// TIA Portal project "Lagerregal_4" (V20) (continued)
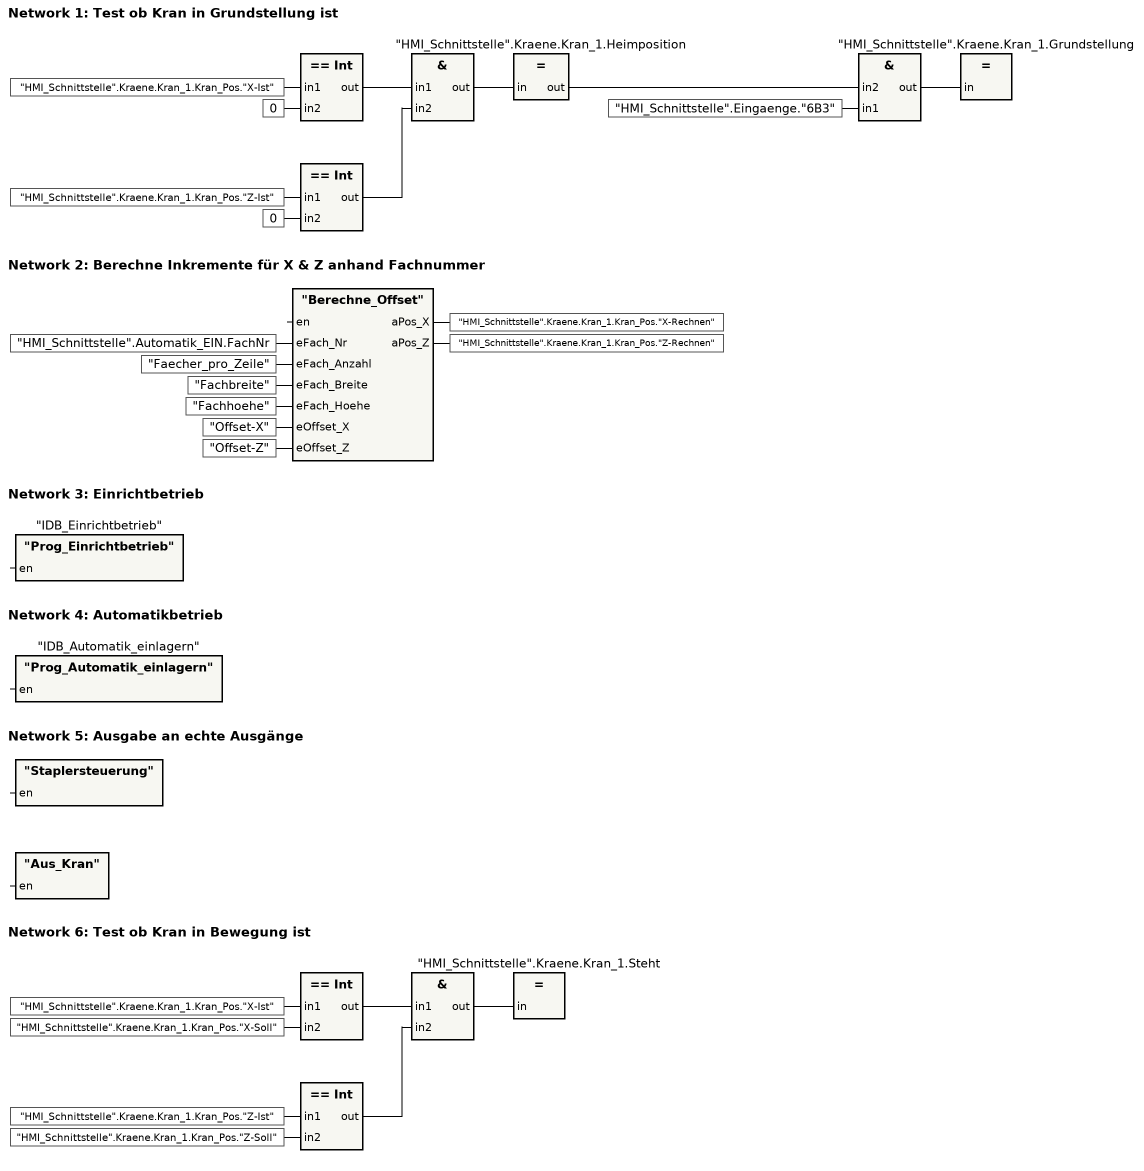
   "HMI_Schnittstelle".Kraene.Kran_1.Heimposition := ("HMI_Schnittstelle".Kraene.Kran_1.Kran_Pos."X-Ist" = 0) AND ("HMI_Schnittstelle".Kraene.Kran_1.Kran_Pos."Z-Ist" = 0);
   "HMI_Schnittstelle".Kraene.Kran_1.Grundstellung := "HMI_Schnittstelle".Kraene.Kran_1.Heimposition AND "HMI_Schnittstelle".Eingaenge."6B3";
END_REGION

REGION Network 2: Berechne Inkremente für X & Z anhand Fachnummer
   "Berechne_Offset"(eFach_Nr := "HMI_Schnittstelle".Automatik_EIN.FachNr,
                     eFach_Anzahl := "Faecher_pro_Zeile",
                     eFach_Breite := "Fachbreite",
                     eFach_Hoehe := "Fachhoehe",
                     eOffset_X := "Offset-X",
                     eOffset_Z := "Offset-Z",
                     aPos_X => "HMI_Schnittstelle".Kraene.Kran_1.Kran_Pos."X-Rechnen",
                     aPos_Z => "HMI_Schnittstelle".Kraene.Kran_1.Kran_Pos."Z-Rechnen");
END_REGION

REGION Network 3: Einrichtbetrieb
   "IDB_Einrichtbetrieb"();   // "Prog_Einrichtbetrieb"
END_REGION

REGION Network 4: Automatikbetrieb
   "IDB_Automatik_einlagern"();   // "Prog_Automatik_einlagern"
END_REGION

REGION Network 5: Ausgabe an echte Ausgänge
   "Staplersteuerung"();
   "Aus_Kran"();
END_REGION

REGION Network 6: Test ob Kran in Bewegung ist
   "HMI_Schnittstelle".Kraene.Kran_1.Steht := ("HMI_Schnittstelle".Kraene.Kran_1.Kran_Pos."X-Ist" = "HMI_Schnittstelle".Kraene.Kran_1.Kran_Pos."X-Soll") AND ("HMI_Schnittstelle".Kraene.Kran_1.Kran_Pos."Z-Ist" = "HMI_Schnittstelle".Kraene.Kran_1.Kran_Pos."Z-Soll");
END_REGION
END_ORGANIZATION_BLOCK

// folder: Bandsteuerung

FUNCTION_BLOCK "Ein_Baender"   // FB20, FBD
{ S7_Optimized_Access := 'TRUE' }
VERSION : 0.1
BEGIN

REGION Network 1 (SCL): Sensoren Einlass
   "HMI_Schnittstelle".Eingaenge."1B1" := NOT "1B1";
   "HMI_Schnittstelle".Eingaenge."1B2" := NOT "1B2";
   "HMI_Schnittstelle".Eingaenge."2B1" := NOT "2B1";
   "HMI_Schnittstelle".Eingaenge."2B2" := NOT "2B2";
   "HMI_Schnittstelle".Eingaenge."3B1" := NOT "3B1";
END_REGION

REGION Network 2 (SCL): Sensoren Auslass
   "HMI_Schnittstelle".Eingaenge."4B1" := NOT "4B1";
   "HMI_Schnittstelle".Eingaenge."5B1" := NOT "5B1";
END_REGION
END_FUNCTION_BLOCK

FUNCTION_BLOCK "Bandsteuerung"   // FB21, FBD
{ S7_Optimized_Access := 'TRUE' }
VERSION : 0.1
   VAR
      RTRIG_Palette_geladen : R_TRIG;
      FTRIG_MDB_1B2 : F_TRIG;
      FTRIG_MDB_2B1 : F_TRIG;
      FTRIG_MDB_2B2 : F_TRIG;
      FTRIG_MDB_5B1 : F_TRIG;
      Band_belegt : Bool;
   END_VAR
BEGIN

REGION Network 1 (SCL): Flankenabfragen
   #RTRIG_Palette_geladen(CLK:="HMI_Schnittstelle".Automatik_EIN.Schrittnummer = 5);
   #FTRIG_MDB_1B2(CLK:="HMI_Schnittstelle".Eingaenge."1B2");
   #FTRIG_MDB_2B1(CLK := "HMI_Schnittstelle".Eingaenge."2B1");
   #FTRIG_MDB_2B2(CLK := "HMI_Schnittstelle".Eingaenge."2B2");
   #FTRIG_MDB_5B1(CLK := "HMI_Schnittstelle".Eingaenge."5B1");
END_REGION

REGION Network 2: Einlasssteuerung
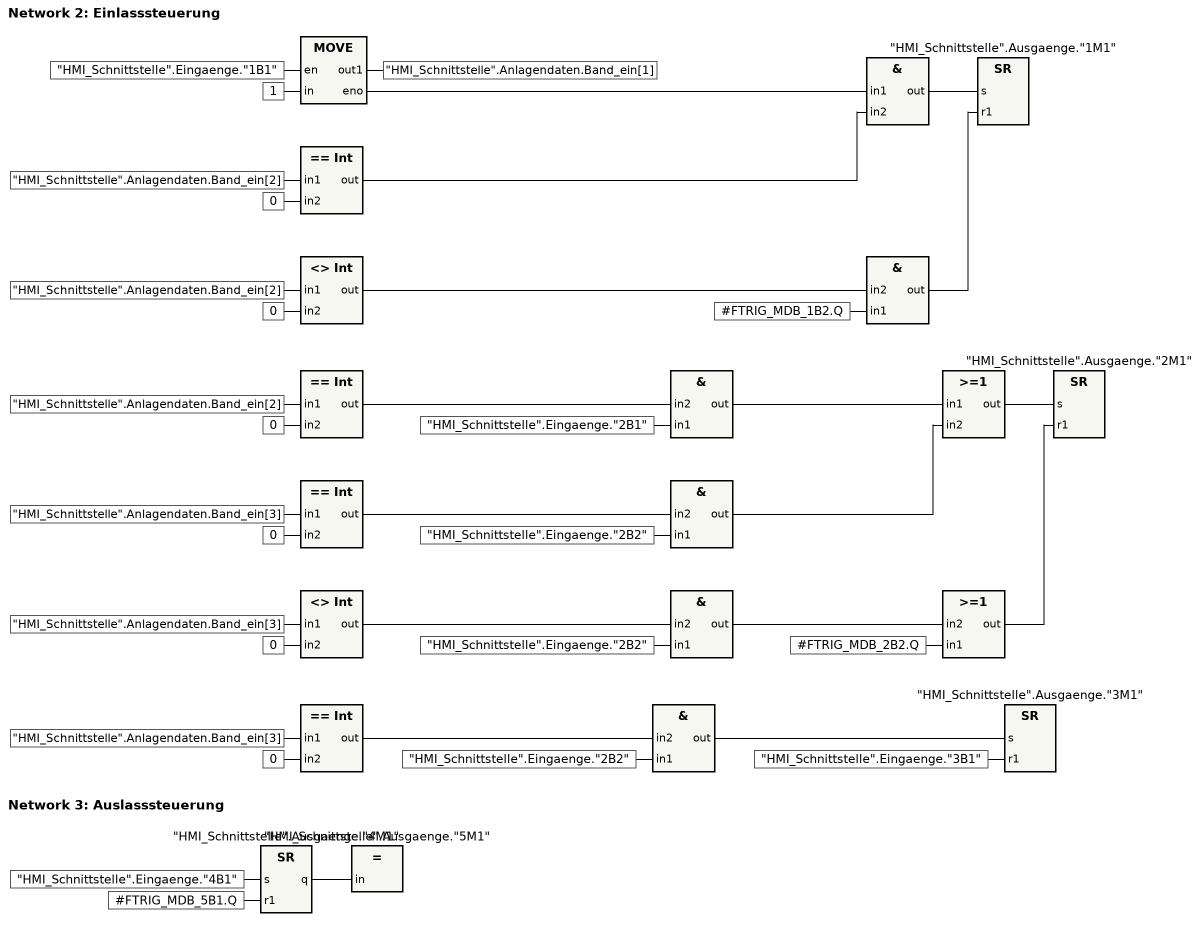
   IF "HMI_Schnittstelle".Eingaenge."1B1" THEN "HMI_Schnittstelle".Anlagendaten.Band_ein[1] := 1; END_IF;
   IF "HMI_Schnittstelle".Eingaenge."1B1" AND ("HMI_Schnittstelle".Anlagendaten.Band_ein[2] = 0) THEN
       "HMI_Schnittstelle".Ausgaenge."1M1" := TRUE;   // SR flip-flop
   END_IF;
   IF ("HMI_Schnittstelle".Anlagendaten.Band_ein[2] <> 0) AND #FTRIG_MDB_1B2.Q THEN
       "HMI_Schnittstelle".Ausgaenge."1M1" := FALSE;
   END_IF;
   IF (("HMI_Schnittstelle".Anlagendaten.Band_ein[2] = 0) AND "HMI_Schnittstelle".Eingaenge."2B1") OR (("HMI_Schnittstelle".Anlagendaten.Band_ein[3] = 0) AND "HMI_Schnittstelle".Eingaenge."2B2") THEN
       "HMI_Schnittstelle".Ausgaenge."2M1" := TRUE;   // SR flip-flop
   END_IF;
   IF (("HMI_Schnittstelle".Anlagendaten.Band_ein[3] <> 0) AND "HMI_Schnittstelle".Eingaenge."2B2") OR #FTRIG_MDB_2B2.Q THEN
       "HMI_Schnittstelle".Ausgaenge."2M1" := FALSE;
   END_IF;
   IF ("HMI_Schnittstelle".Anlagendaten.Band_ein[3] = 0) AND "HMI_Schnittstelle".Eingaenge."2B2" THEN
       "HMI_Schnittstelle".Ausgaenge."3M1" := TRUE;   // SR flip-flop
   END_IF;
   IF "HMI_Schnittstelle".Eingaenge."3B1" THEN "HMI_Schnittstelle".Ausgaenge."3M1" := FALSE; END_IF;
END_REGION

REGION Network 3: Auslasssteuerung
   IF "HMI_Schnittstelle".Eingaenge."4B1" THEN
       "HMI_Schnittstelle".Ausgaenge."4M1" := TRUE;   // SR flip-flop
   END_IF;
   IF #FTRIG_MDB_5B1.Q THEN "HMI_Schnittstelle".Ausgaenge."4M1" := FALSE; END_IF;
   "HMI_Schnittstelle".Ausgaenge."5M1" := "HMI_Schnittstelle".Ausgaenge."4M1";
END_REGION

REGION Network 4 (SCL): Bandbelegung
   IF #FTRIG_MDB_2B1.Q THEN
       "HMI_Schnittstelle".Anlagendaten.Band_ein[2] := "HMI_Schnittstelle".Anlagendaten.Band_ein[1];
       "HMI_Schnittstelle".Anlagendaten.Band_ein[1] := 0;
   END_IF;

   IF #FTRIG_MDB_2B2.Q THEN
       "HMI_Schnittstelle".Anlagendaten.Band_ein[3] := "HMI_Schnittstelle".Anlagendaten.Band_ein[2];
       "HMI_Schnittstelle".Anlagendaten.Band_ein[2] := 0;
   END_IF;

   IF #RTRIG_Palette_geladen.Q THEN
       "HMI_Schnittstelle".Anlagendaten.Band_ein[3] := 0;
   END_IF;
END_REGION
END_FUNCTION_BLOCK

FUNCTION "Aus_Baender" : Void   // FC20, FBD
{ S7_Optimized_Access := 'TRUE' }
VERSION : 0.1
BEGIN

REGION Network 1 (SCL): Bänder Einlass
   "1M1" := "HMI_Schnittstelle".Ausgaenge."1M1";
   "2M1" := "HMI_Schnittstelle".Ausgaenge."2M1";
   "3M1" := "HMI_Schnittstelle".Ausgaenge."3M1";
END_REGION

REGION Network 2 (SCL): Bänder Auslass
   "4M1" := "HMI_Schnittstelle".Ausgaenge."4M1";
   "5M1" := "HMI_Schnittstelle".Ausgaenge."5M1";
END_REGION
END_FUNCTION

ORGANIZATION_BLOCK "Main_Baender"   // OB124, FBD, ProgramCycle
TITLE = "Main Program Sweep (Cycle)"
{ S7_Optimized_Access := 'TRUE' }
VERSION : 0.1
   VAR_INPUT
      Initial_Call : Bool;   // Initial call of this OB
      Remanence : Bool;   // =True, if remanent data are available
   END_VAR
BEGIN

REGION Network 1
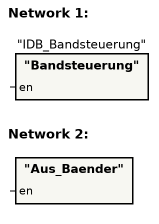
   "IDB_Bandsteuerung"();   // "Bandsteuerung"
END_REGION

REGION Network 2
   "Aus_Baender"();
END_REGION
END_ORGANIZATION_BLOCK

// folder: HMI

FUNCTION_BLOCK "Prog_Einrichtbetrieb"   // FB3, FBD
{ S7_Optimized_Access := 'TRUE' }
VERSION : 0.1
   VAR
      "PTRIG_MDB_X-Pos" : R_TRIG;
      "PTRIG_MDB_X-Neg" : R_TRIG;
      "PTRIG_MDB_Z-Pos" : R_TRIG;
      "PTRIG_MDB_Z-Neg" : R_TRIG;
   END_VAR
BEGIN

REGION Network 1: Button Flanken erfassen
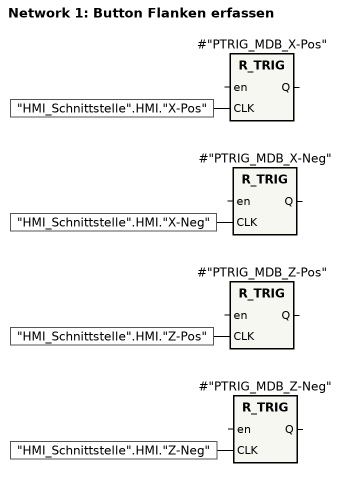
   #"PTRIG_MDB_X-Pos"(CLK := "HMI_Schnittstelle".HMI."X-Pos");   // R_TRIG
   #"PTRIG_MDB_X-Neg"(CLK := "HMI_Schnittstelle".HMI."X-Neg");   // R_TRIG
   #"PTRIG_MDB_Z-Pos"(CLK := "HMI_Schnittstelle".HMI."Z-Pos");   // R_TRIG
   #"PTRIG_MDB_Z-Neg"(CLK := "HMI_Schnittstelle".HMI."Z-Neg");   // R_TRIG
END_REGION

REGION Network 2 (SCL): Achsen inkrementieren
   // X-Achse Inkrementieren
   IF #"PTRIG_MDB_X-Pos".Q THEN
       "HMI_Schnittstelle".Kraene.Kran_1.Kran_Pos."X-Soll" += UINT_TO_INT("HMI_Schnittstelle".HMI.Inkrement);
   END_IF;

   IF #"PTRIG_MDB_X-Neg".Q THEN
       "HMI_Schnittstelle".Kraene.Kran_1.Kran_Pos."X-Soll" -= UINT_TO_INT("HMI_Schnittstelle".HMI.Inkrement);
   END_IF;


   // Z-Achse Inkrementieren
   IF #"PTRIG_MDB_Z-Pos".Q THEN
       "HMI_Schnittstelle".Kraene.Kran_1.Kran_Pos."Z-Soll" += UINT_TO_INT("HMI_Schnittstelle".HMI.Inkrement);
   END_IF;

   IF #"PTRIG_MDB_Z-Neg".Q THEN
       "HMI_Schnittstelle".Kraene.Kran_1.Kran_Pos."Z-Soll" -= UINT_TO_INT("HMI_Schnittstelle".HMI.Inkrement);
   END_IF;
END_REGION
END_FUNCTION_BLOCK

FUNCTION_BLOCK "Ein_HMI"   // FB10, FBD
{ S7_Optimized_Access := 'TRUE' }
VERSION : 0.1
BEGIN
END_FUNCTION_BLOCK

// folder: Kransteuerung

FUNCTION_BLOCK "FC_Kran_beladen"   // FB25, FBD
{ S7_Optimized_Access := 'TRUE' }
VERSION : 0.1
   VAR_INPUT
      "eKran_Z-Ist" : Int;
      eSchrittnummer : Int;
   END_VAR
   VAR_OUTPUT
      aGabel : Bool;
      aBeladen : Bool;
      "aKran_Z-Soll" : Int;
   END_VAR
   VAR
      PTRIG_Schritt2 : Bool;
   END_VAR
   VAR_TEMP   // added for the SCL form of the ladder/FBD networks
      _w1 : Bool;
      _w2 : Bool;
   END_VAR
BEGIN

REGION Network 1: Gabel zur Seite ausfahren
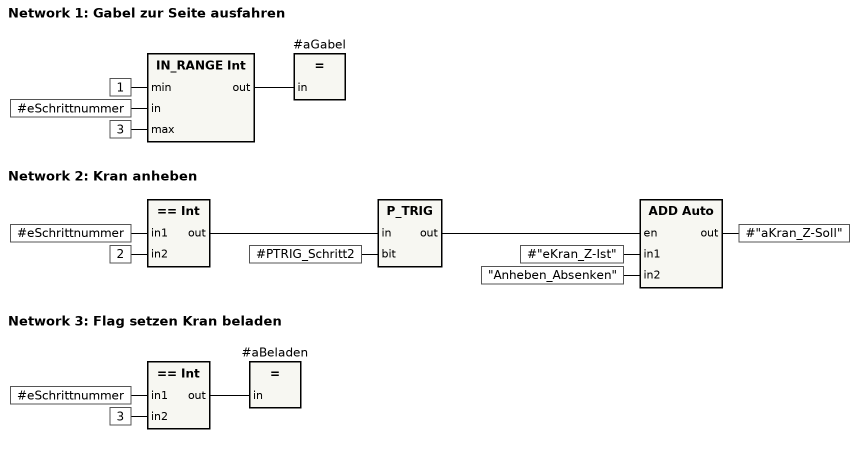
   #aGabel := (1 <= #eSchrittnummer) AND (#eSchrittnummer <= 3);
END_REGION

REGION Network 2: Kran anheben
   #_w1 := #eSchrittnummer = 2;
   #_w2 := #_w1 AND NOT #PTRIG_Schritt2;   // rising edge
   #PTRIG_Schritt2 := #_w1;
   IF #_w2 THEN #"aKran_Z-Soll" := #"eKran_Z-Ist" + "Anheben_Absenken"; END_IF;
END_REGION

REGION Network 3: Flag setzen Kran beladen
   #aBeladen := #eSchrittnummer = 3;
END_REGION
END_FUNCTION_BLOCK

FUNCTION_BLOCK "FC_Kran_entladen"   // FB26, FBD
{ S7_Optimized_Access := 'TRUE' }
VERSION : 0.1
   VAR_INPUT
      "eKran_Z-Ist" : Int;
      eSchrittnummer : Int;
   END_VAR
   VAR_OUTPUT
      aGabel : Bool;
      aBeladen : Bool;
      "aKran_Z-Soll" : Int;
   END_VAR
   VAR
      PTRIG_Schritt2 : Bool;
   END_VAR
   VAR_TEMP   // added for the SCL form of the ladder/FBD networks
      _w1 : Bool;
      _w2 : Bool;
   END_VAR
BEGIN

REGION Network 1: Gabel zur Seite ausfahren
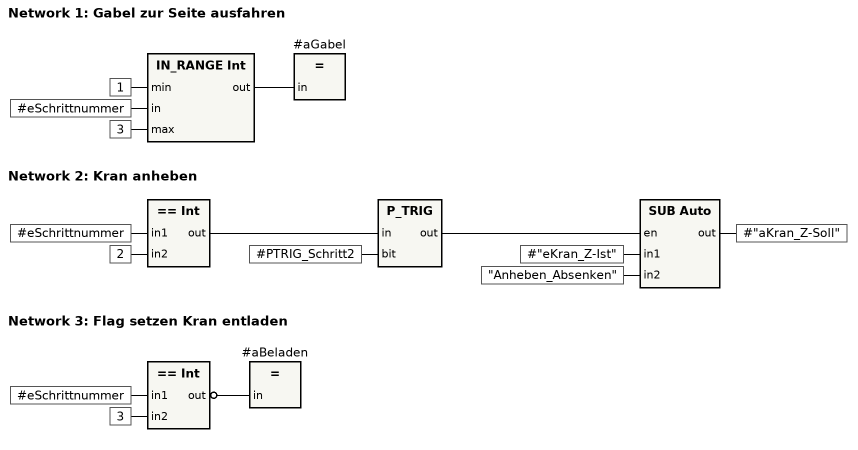
   #aGabel := (1 <= #eSchrittnummer) AND (#eSchrittnummer <= 3);
END_REGION

REGION Network 2: Kran anheben
   #_w1 := #eSchrittnummer = 2;
   #_w2 := #_w1 AND NOT #PTRIG_Schritt2;   // rising edge
   #PTRIG_Schritt2 := #_w1;
   IF #_w2 THEN #"aKran_Z-Soll" := #"eKran_Z-Ist" - "Anheben_Absenken"; END_IF;
END_REGION

REGION Network 3: Flag setzen Kran entladen
   #aBeladen := NOT (#eSchrittnummer = 3);
END_REGION
END_FUNCTION_BLOCK

FUNCTION_BLOCK "Ein_Kran"   // FB30, FBD
{ S7_Optimized_Access := 'TRUE' }
VERSION : 0.1
   VAR
      NTRIG_MDB_1B2 : F_TRIG;
      NTRIG_MDB_2B2 : F_TRIG;
      NTRIG_MDB_5B1 : F_TRIG;
   END_VAR
BEGIN

REGION Network 1 (SCL): Sensoren Kran_1
   "HMI_Schnittstelle".Eingaenge."6B1" := "6B1";
   "HMI_Schnittstelle".Eingaenge."6B2" := "6B2";
   "HMI_Schnittstelle".Eingaenge."6B3" := "6B3";
END_REGION

REGION Network 2: Kran_1 Position einlesen
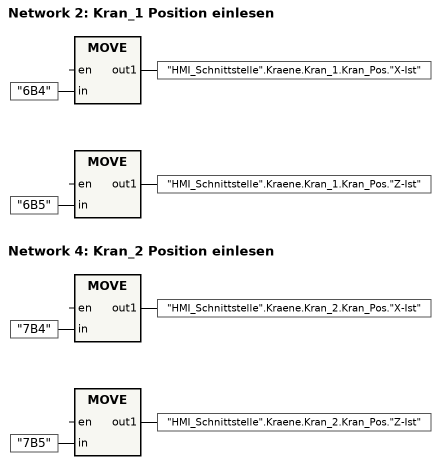
   "HMI_Schnittstelle".Kraene.Kran_1.Kran_Pos."X-Ist" := "6B4";
   "HMI_Schnittstelle".Kraene.Kran_1.Kran_Pos."Z-Ist" := "6B5";
END_REGION

REGION Network 3 (SCL): Sensoren Kran_2
   "HMI_Schnittstelle".Eingaenge."7B1" := "7B1";
   "HMI_Schnittstelle".Eingaenge."7B2" := "7B2";
   "HMI_Schnittstelle".Eingaenge."7B3" := "7B3";
END_REGION

REGION Network 4: Kran_2 Position einlesen
   "HMI_Schnittstelle".Kraene.Kran_2.Kran_Pos."X-Ist" := "7B4";
   "HMI_Schnittstelle".Kraene.Kran_2.Kran_Pos."Z-Ist" := "7B5";
END_REGION
END_FUNCTION_BLOCK

FUNCTION "Aus_Kran" : Void   // FC30, FBD
{ S7_Optimized_Access := 'TRUE' }
VERSION : 0.1
BEGIN

REGION Network 1 (SCL): Achsen Kräne Soll-Pos
   // Kran Position
   // Kran X-Soll-Position
   (*
   "6M4" := "HMI_Schnittstelle".Kraene.Kran_1.Kran_Pos."X-Soll";
   "6M5" := "HMI_Schnittstelle".Kraene.Kran_2.Kran_Pos."X-Soll";
   *)

   // Kran Z-Soll-Position
   (*
   "7M4" := "HMI_Schnittstelle".Kraene.Kran_1.Kran_Pos."Z-Soll";
   "7M5" := "HMI_Schnittstelle".Kraene.Kran_2.Kran_Pos."Z-Soll";
   *)
END_REGION

REGION Network 2 (SCL): Kräne Gabelsteuerung
   "6M1" := "HMI_Schnittstelle".Ausgaenge."6M1";
   "6M2" := "HMI_Schnittstelle".Ausgaenge."6M2";

   "7M1" := "HMI_Schnittstelle".Ausgaenge."7M1";
   "7M2" := "HMI_Schnittstelle".Ausgaenge."7M2";
END_REGION
END_FUNCTION

FUNCTION "Staplersteuerung" : Void   // FC70, FBD
{ S7_Optimized_Access := 'TRUE' }
VERSION : 0.1
BEGIN

REGION Network 1: Sollposition X
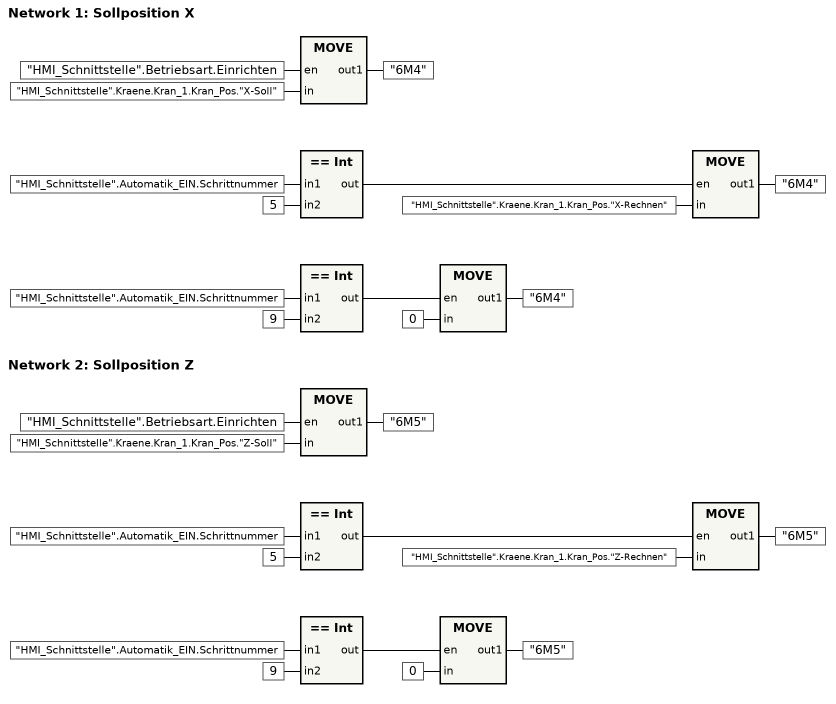
   IF "HMI_Schnittstelle".Betriebsart.Einrichten THEN
       "6M4" := "HMI_Schnittstelle".Kraene.Kran_1.Kran_Pos."X-Soll";
   END_IF;
   IF "HMI_Schnittstelle".Automatik_EIN.Schrittnummer = 5 THEN
       "6M4" := "HMI_Schnittstelle".Kraene.Kran_1.Kran_Pos."X-Rechnen";
   END_IF;
   IF "HMI_Schnittstelle".Automatik_EIN.Schrittnummer = 9 THEN "6M4" := 0; END_IF;
END_REGION

REGION Network 2: Sollposition Z
   IF "HMI_Schnittstelle".Betriebsart.Einrichten THEN
       "6M5" := "HMI_Schnittstelle".Kraene.Kran_1.Kran_Pos."Z-Soll";
   END_IF;
   IF "HMI_Schnittstelle".Automatik_EIN.Schrittnummer = 5 THEN
       "6M5" := "HMI_Schnittstelle".Kraene.Kran_1.Kran_Pos."Z-Rechnen";
   END_IF;
   IF "HMI_Schnittstelle".Automatik_EIN.Schrittnummer = 9 THEN "6M5" := 0; END_IF;
END_REGION

REGION Network 3 (SCL): Z-Achse Kran_1 Soll-Pos
   // Einrichtbetrieb
   IF "HMI_Schnittstelle".Betriebsart.Einrichten THEN
       "6M5" := "HMI_Schnittstelle".Kraene.Kran_1.Kran_Pos."Z-Soll";

   // Automatikbetrieb    
   ELSIF "HMI_Schnittstelle".Automatik_EIN.Schrittnummer = 3 THEN
       // Palette aus Grundstellung anheben
       "6M5" := "Anheben_Absenken" + 2;
   ELSIF "HMI_Schnittstelle".Automatik_EIN.Schrittnummer = 5 THEN
       //Fach mit Nummer anfahren
       "6M5" := "HMI_Schnittstelle".Kraene.Kran_1.Kran_Pos."Z-Rechnen";
   ELSIF "HMI_Schnittstelle".Automatik_EIN.Schrittnummer = 7 THEN
       // Palette in Regal einlagern
       "6M5" := "HMI_Schnittstelle".Kraene.Kran_1.Kran_Pos."Z-Rechnen" - "Anheben_Absenken";
   ELSIF "HMI_Schnittstelle".Automatik_EIN.Schrittnummer = 9 THEN
       // Stapler in Grundstellung
       "6M5" := 0;
   END_IF;
END_REGION

REGION Network 4 (SCL): Gabel links ausfahren
   "HMI_Schnittstelle".Ausgaenge."6M1" := "HMI_Schnittstelle".Automatik_EIN.Schrittnummer = 2
                                       OR "HMI_Schnittstelle".Automatik_EIN.Schrittnummer = 3;
END_REGION

REGION Network 5 (SCL): Gabel rechts ausfahren
   "HMI_Schnittstelle".Ausgaenge."6M2" := "HMI_Schnittstelle".Automatik_EIN.Schrittnummer = 6
                                       OR "HMI_Schnittstelle".Automatik_EIN.Schrittnummer = 7;
END_REGION
END_FUNCTION

(* ===== HMI "HMI_RT_1" =====
system functions are stored by id; their names below are inferred from use
connection "HMI_Verbindung_1": ETHERNET, S7_1500_OMS

HMI tags "Standard-Variablentabelle"
   "HMI_Schnittstelle_Kraene_Kran_1_Z-Soll" : Int = PLC HMI_Schnittstelle.Kraene.Kran_1.Kran_Pos.Z-Soll, 100 ms
   "HMI_Schnittstelle_Kraene_Kran_1_X-Soll" : Int = PLC HMI_Schnittstelle.Kraene.Kran_1.Kran_Pos.X-Soll, 100 ms
   "HMI_Schnittstelle_Kraene_Kran_1_X-Ist" : Int = PLC HMI_Schnittstelle.Kraene.Kran_1.Kran_Pos.X-Ist, 100 ms
   "HMI_Schnittstelle_Kraene_Kran_1_Z-Ist" : Int = PLC HMI_Schnittstelle.Kraene.Kran_1.Kran_Pos.Z-Ist, 100 ms
   "HMI_Schnittstelle_HMI_X-Neg" : Bool = PLC HMI_Schnittstelle.HMI.X-Neg, 1 s
   "HMI_Schnittstelle_HMI_X-Pos" : Bool = PLC HMI_Schnittstelle.HMI.X-Pos, 1 s
   "HMI_Schnittstelle_HMI_Z-Neg" : Bool = PLC HMI_Schnittstelle.HMI.Z-Neg, 1 s
   "HMI_Schnittstelle_HMI_Z-Pos" : Bool = PLC HMI_Schnittstelle.HMI.Z-Pos, 1 s
   "HMI_Schnittstelle_HMI_Inkrement" : UInt = PLC HMI_Schnittstelle.HMI.Inkrement, 1 s
   "HMI_Schnittstelle_Ausgaenge_Fach_ansteuern" : Bool = PLC HMI_Schnittstelle.Fach_ansteuern, 1 s
   "HMI_Schnittstelle_Ausgaenge_Fach" : Int = PLC HMI_Schnittstelle.Fach, 1 s
   "Clock_1Hz" : Bool = PLC Clock_1Hz AT %M0.5, 100 ms
   "HMI_Schnittstelle_Fach" : Int = PLC HMI_Schnittstelle.Fach, 1 s
   "HMI_Schnittstelle_Fach_ansteuern" : Bool = PLC HMI_Schnittstelle.Fach_ansteuern, 1 s
   "Warenlager_Lager{1}_Flags_Belegt" : Bool = PLC Warenlager.Lager[1].Flags.Belegt, 1 s
   "Warenlager_Lager{1}_Flags_In_Benutzung" : Bool = PLC Warenlager.Lager[1].Flags.In_Benutzung, 1 s
   "HMI_Schnittstelle_Automatik_EIN_FachNr" : Int = PLC HMI_Schnittstelle.Automatik_EIN.FachNr, 500 ms

HMI tags "Interne_Variablen"
   "Bildnummer" : Int, internal

text list "Liste_Bilder": 0..1 'Bitte Bild auswählen'; 1 'Startbild'; 2 'Betriebsart'; 3 'Handbetrieb'; 4 ''; 5 'Einrichtbetrieb'; 6 'Statistik'; 7 ''; 8 'Meldungen'; 9 'Diagnose'; 10 'Benutzerverwaltung'

screen "01_Lageransicht" 800x420, template "Menüleiste"
   on GenerateScreen: SetTag("Bildnummer", 1)
   Button "Schaltfläche_4" at 10,438 size 96x32; TextOff 'Teachen'
      on Press: ActivateScreen("05_Teachmodus", 0)
   Rectangle "Rechteck_1" at 650,280 size 50x50
      Appearance <- "Warenlager_Lager{1}_Flags_Belegt"
   TextField "Textfeld_1" at 650,280 size 50x50; Text '1'
      Appearance <- "Warenlager_Lager{1}_Flags_In_Benutzung"

screen "05_Teachmodus" 800x420, template "Menüleiste"
   on GenerateScreen: SetTag("Bildnummer", 5)
   Button "Schaltfläche_1" at 694,10 size 96x32; TextOff 'Zurück'
      on Press: function_efd93a16()
   TextField "Textfeld_1" at 308,10 size 184x23; Text 'Kalibrierungsmodus'
   Slider "Schieberegler_2" at 113,300 size 230x50; Caption 'Breite'
      ProcessValue <- "HMI_Schnittstelle_Kraene_Kran_1_X-Soll"
   IOField "EA-Feld_8" at 370,67 size 96x32; FormatPattern 99999
      ProcessValue <- "HMI_Schnittstelle_Kraene_Kran_1_X-Ist"
   IOField "EA-Feld_9" at 485,68 size 96x32; FormatPattern 99999
      ProcessValue <- "HMI_Schnittstelle_Kraene_Kran_1_Z-Ist"
   Slider "Schieberegler_1" at 10,37 size 50x230; Caption 'Höhe'
      ProcessValue <- "HMI_Schnittstelle_Kraene_Kran_1_Z-Soll"
   Button "Schaltfläche_5" at 345,300 size 25x50; TextOff '-'
      on Press: function_b14e0dd5("HMI_Schnittstelle_HMI_X-Neg", 0)
      Appearance <- "HMI_Schnittstelle_HMI_X-Neg"
   IOField "EA-Feld_7" at 10,300 size 70x50; FormatPattern 99999
      ProcessValue <- "HMI_Schnittstelle_HMI_Inkrement"
   Button "Schaltfläche_7" at 10,269 size 50x25; TextOff '-'
      on Press: function_b14e0dd5("HMI_Schnittstelle_HMI_Z-Neg", 0)
      Appearance <- "HMI_Schnittstelle_HMI_Z-Neg"
   Button "Schaltfläche_8" at 10,10 size 50x25; TextOff '+'
      on Press: function_b14e0dd5("HMI_Schnittstelle_HMI_Z-Pos", 0)
      Appearance <- "HMI_Schnittstelle_HMI_Z-Pos"
   Button "Schaltfläche_6" at 86,300 size 25x50; TextOff '+'
      on Press: function_b14e0dd5("HMI_Schnittstelle_HMI_X-Pos", 0)
      Appearance <- "HMI_Schnittstelle_HMI_X-Pos"
   TextField "Textfeld_2" at 370,42 size 111x23; Text 'Ist-X-Achse'
   TextField "Textfeld_3" at 485,42 size 110x23; Text 'Ist-Z-Achse'
   TextField "Textfeld_4" at 370,103 size 88x23; Text 'Fach-Nr.:'
   IOField "EA-Feld_1" at 370,128 size 96x32; FormatPattern 99
      ProcessValue <- "HMI_Schnittstelle_Fach"
   Button "Schaltfläche_2" at 485,128 size 96x32; TextOff 'Testen'
      on Press: function_b14e0dd5("HMI_Schnittstelle_Fach_ansteuern", 0)

screen "Detailansicht" 800x420, template "Menüleiste"
   Button "Schaltfläche_1" at 694,10 size 96x32; TextOff 'Zurück'
      on Press: function_efd93a16()

Template "Menüleiste" 800x420
   Button "Vorlage_Schaltfläche_1" at 0,360 size 80x60; TextOff 'HOME'; PictureOff "Grafik_2"; PictureOn "Grafik_2"
      Appearance <- "Bildnummer"
      on Press: ActivateScreen("01_Lageransicht", 0)
   Button "Vorlage_Schaltfläche_2" at 80,360 size 80x60; TextOff 'BETRIEB'; PictureOff "Grafik_8"; PictureOn "Grafik_8"
      Appearance <- "Bildnummer"
      on Press: ActivateScreen("02_Bild", 0)
   Button "Vorlage_Schaltfläche_3" at 160,360 size 80x60; TextOff 'HAND'; PictureOff "Grafik_7"; PictureOn "Grafik_7"
      Appearance <- "Bildnummer"
      on Press: ActivateScreen("03_Bild", 0)
   Button "Vorlage_Schaltfläche_4" at 240,360 size 80x60; TextOff 'Text'
      Appearance <- "Bildnummer"
      on Press: ActivateScreen("04_Bild", 0)
   Button "Vorlage_Schaltfläche_5" at 320,360 size 80x60; TextOff 'TEACH'; PictureOn "Grafik_3"; PictureOff "Grafik_3"; Authorization "Einstellen"
      Appearance <- "Bildnummer"
      on Press: ActivateScreen("05_Teachmodus", 0)
   Button "Vorlage_Schaltfläche_6" at 400,360 size 80x60; TextOff 'STATS'; PictureOff "Grafik_4"; PictureOn "Grafik_4"
      Appearance <- "Bildnummer"
      on Press: ActivateScreen("06_Statistik", 0)
   Button "Vorlage_Schaltfläche_7" at 480,360 size 80x60; TextOff 'Text'
      Appearance <- "Bildnummer"
      on Press: ActivateScreen("07_Bild", 0)
   Button "Vorlage_Schaltfläche_8" at 560,360 size 80x60; TextOff 'FEHLER'; PictureOff "Grafik_6"; PictureOn "Grafik_6"
      Appearance <- "Bildnummer"
      on Press: ActivateScreen("08_Bild", 0)
   Button "Vorlage_Schaltfläche_9" at 640,360 size 80x60; TextOff 'DIAG'; PictureOff "Grafik_9"; PictureOn "Grafik_9"
      Appearance <- "Bildnummer"
      on Press: ActivateScreen("09_Diagnose", 0)
   Button "Vorlage_Schaltfläche_10" at 720,360 size 80x60; TextOff 'NUTZER'; PictureOff "Grafik_10"; PictureOn "Grafik_10"
      Appearance <- "Bildnummer"
      on Press: ActivateScreen("10_Benutzer", 0)

screen "02_Bild" 800x420, template "Menüleiste"
   on GenerateScreen: SetTag("Bildnummer", 2)

screen "03_Bild" 800x420, template "Menüleiste"
   on GenerateScreen: SetTag("Bildnummer", 3)

screen "04_Bild" 800x420, template "Menüleiste"
   on GenerateScreen: SetTag("Bildnummer", 4)

screen "06_Statistik" 800x420, template "Menüleiste"
   on GenerateScreen: SetTag("Bildnummer", 6)
   TrendView "Kurvenanzeige_1" at 10,10 size 780x340

screen "07_Bild" 800x420, template "Menüleiste"
   on GenerateScreen: SetTag("Bildnummer", 7)

screen "08_Bild" 800x420, template "Menüleiste"
   on GenerateScreen: SetTag("Bildnummer", 8)

screen "09_Diagnose" 800x420, template "Menüleiste"
   on GenerateScreen: SetTag("Bildnummer", 9)
   SysDiagControl "System-Diagnoseanzeige_1" at 10,10 size 780x340

screen "10_Benutzer" 800x420, template "Menüleiste"
   on GenerateScreen: SetTag("Bildnummer", 10)
   UserView "Benutzeranzeige_1" at 10,10 size 780x340
*)